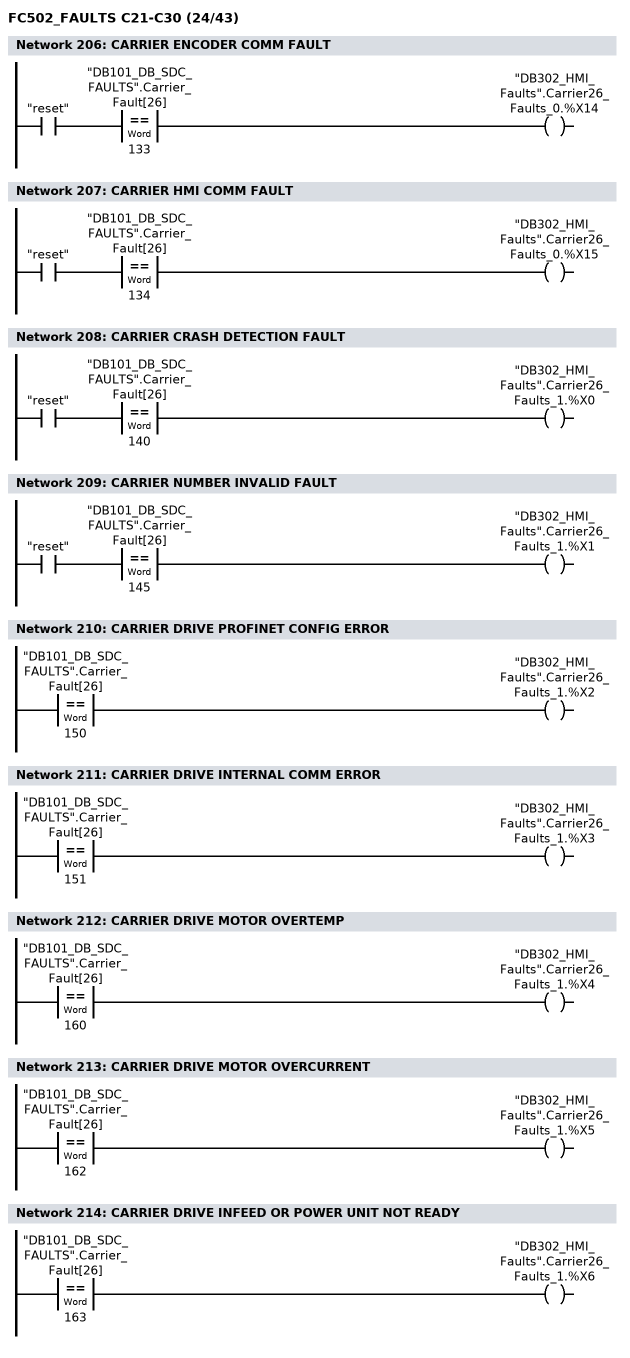
   RUNG wire#powerrail
      Contact( "reset" )
      { S7_Templates := "SrcType := Word" } EQ_Contact(in1 := "DB101_DB_SDC_FAULTS".Carrier_Fault[26], in2 := 133)
      Coil( "DB302_HMI_Faults".Carrier26_Faults_0.%X14 )
   END_RUNG
   // the same network as SCL:
   "DB302_HMI_Faults".Carrier26_Faults_0.%X14 := "reset" AND ("DB101_DB_SDC_FAULTS".Carrier_Fault[26] = 133);
END_REGION

REGION Network 207: CARRIER HMI COMM FAULT
   RUNG wire#powerrail
      Contact( "reset" )
      { S7_Templates := "SrcType := Word" } EQ_Contact(in1 := "DB101_DB_SDC_FAULTS".Carrier_Fault[26], in2 := 134)
      Coil( "DB302_HMI_Faults".Carrier26_Faults_0.%X15 )
   END_RUNG
   // the same network as SCL:
   "DB302_HMI_Faults".Carrier26_Faults_0.%X15 := "reset" AND ("DB101_DB_SDC_FAULTS".Carrier_Fault[26] = 134);
END_REGION

REGION Network 208: CARRIER CRASH DETECTION FAULT
   RUNG wire#powerrail
      Contact( "reset" )
      { S7_Templates := "SrcType := Word" } EQ_Contact(in1 := "DB101_DB_SDC_FAULTS".Carrier_Fault[26], in2 := 140)
      Coil( "DB302_HMI_Faults".Carrier26_Faults_1.%X0 )
   END_RUNG
   // the same network as SCL:
   "DB302_HMI_Faults".Carrier26_Faults_1.%X0 := "reset" AND ("DB101_DB_SDC_FAULTS".Carrier_Fault[26] = 140);
END_REGION

REGION Network 209: CARRIER NUMBER INVALID FAULT
   RUNG wire#powerrail
      Contact( "reset" )
      { S7_Templates := "SrcType := Word" } EQ_Contact(in1 := "DB101_DB_SDC_FAULTS".Carrier_Fault[26], in2 := 145)
      Coil( "DB302_HMI_Faults".Carrier26_Faults_1.%X1 )
   END_RUNG
   // the same network as SCL:
   "DB302_HMI_Faults".Carrier26_Faults_1.%X1 := "reset" AND ("DB101_DB_SDC_FAULTS".Carrier_Fault[26] = 145);
END_REGION

REGION Network 210: CARRIER DRIVE PROFINET CONFIG ERROR
   RUNG wire#powerrail
      { S7_Templates := "SrcType := Word" } EQ_Contact(in1 := "DB101_DB_SDC_FAULTS".Carrier_Fault[26], in2 := 150)
      Coil( "DB302_HMI_Faults".Carrier26_Faults_1.%X2 )
   END_RUNG
   // the same network as SCL:
   "DB302_HMI_Faults".Carrier26_Faults_1.%X2 := "DB101_DB_SDC_FAULTS".Carrier_Fault[26] = 150;
END_REGION

REGION Network 211: CARRIER DRIVE INTERNAL COMM ERROR
   RUNG wire#powerrail
      { S7_Templates := "SrcType := Word" } EQ_Contact(in1 := "DB101_DB_SDC_FAULTS".Carrier_Fault[26], in2 := 151)
      Coil( "DB302_HMI_Faults".Carrier26_Faults_1.%X3 )
   END_RUNG
   // the same network as SCL:
   "DB302_HMI_Faults".Carrier26_Faults_1.%X3 := "DB101_DB_SDC_FAULTS".Carrier_Fault[26] = 151;
END_REGION

REGION Network 212: CARRIER DRIVE MOTOR OVERTEMP
   RUNG wire#powerrail
      { S7_Templates := "SrcType := Word" } EQ_Contact(in1 := "DB101_DB_SDC_FAULTS".Carrier_Fault[26], in2 := 160)
      Coil( "DB302_HMI_Faults".Carrier26_Faults_1.%X4 )
   END_RUNG
   // the same network as SCL:
   "DB302_HMI_Faults".Carrier26_Faults_1.%X4 := "DB101_DB_SDC_FAULTS".Carrier_Fault[26] = 160;
END_REGION

REGION Network 213: CARRIER DRIVE MOTOR OVERCURRENT
   RUNG wire#powerrail
      { S7_Templates := "SrcType := Word" } EQ_Contact(in1 := "DB101_DB_SDC_FAULTS".Carrier_Fault[26], in2 := 162)
      Coil( "DB302_HMI_Faults".Carrier26_Faults_1.%X5 )
   END_RUNG
   // the same network as SCL:
   "DB302_HMI_Faults".Carrier26_Faults_1.%X5 := "DB101_DB_SDC_FAULTS".Carrier_Fault[26] = 162;
END_REGION

REGION Network 214: CARRIER DRIVE INFEED OR POWER UNIT NOT READY
   RUNG wire#powerrail
      { S7_Templates := "SrcType := Word" } EQ_Contact(in1 := "DB101_DB_SDC_FAULTS".Carrier_Fault[26], in2 := 163)
      Coil( "DB302_HMI_Faults".Carrier26_Faults_1.%X6 )
   END_RUNG
   // the same network as SCL:
   "DB302_HMI_Faults".Carrier26_Faults_1.%X6 := "DB101_DB_SDC_FAULTS".Carrier_Fault[26] = 163;
END_REGION

REGION Network 215: CARRIER DRIVE SHORT CIRCUIT / GROUND FAULT DETECTED
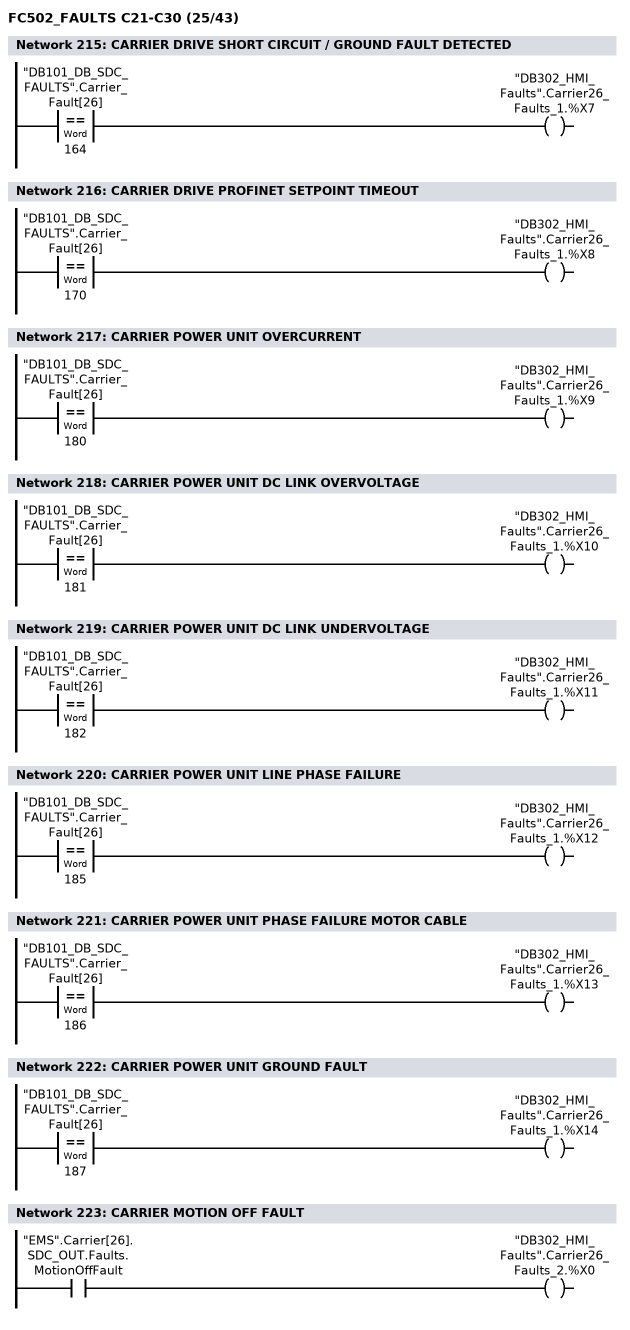
   RUNG wire#powerrail
      { S7_Templates := "SrcType := Word" } EQ_Contact(in1 := "DB101_DB_SDC_FAULTS".Carrier_Fault[26], in2 := 164)
      Coil( "DB302_HMI_Faults".Carrier26_Faults_1.%X7 )
   END_RUNG
   // the same network as SCL:
   "DB302_HMI_Faults".Carrier26_Faults_1.%X7 := "DB101_DB_SDC_FAULTS".Carrier_Fault[26] = 164;
END_REGION

REGION Network 216: CARRIER DRIVE PROFINET SETPOINT TIMEOUT
   RUNG wire#powerrail
      { S7_Templates := "SrcType := Word" } EQ_Contact(in1 := "DB101_DB_SDC_FAULTS".Carrier_Fault[26], in2 := 170)
      Coil( "DB302_HMI_Faults".Carrier26_Faults_1.%X8 )
   END_RUNG
   // the same network as SCL:
   "DB302_HMI_Faults".Carrier26_Faults_1.%X8 := "DB101_DB_SDC_FAULTS".Carrier_Fault[26] = 170;
END_REGION

REGION Network 217: CARRIER POWER UNIT OVERCURRENT
   RUNG wire#powerrail
      { S7_Templates := "SrcType := Word" } EQ_Contact(in1 := "DB101_DB_SDC_FAULTS".Carrier_Fault[26], in2 := 180)
      Coil( "DB302_HMI_Faults".Carrier26_Faults_1.%X9 )
   END_RUNG
   // the same network as SCL:
   "DB302_HMI_Faults".Carrier26_Faults_1.%X9 := "DB101_DB_SDC_FAULTS".Carrier_Fault[26] = 180;
END_REGION

REGION Network 218: CARRIER POWER UNIT DC LINK OVERVOLTAGE
   RUNG wire#powerrail
      { S7_Templates := "SrcType := Word" } EQ_Contact(in1 := "DB101_DB_SDC_FAULTS".Carrier_Fault[26], in2 := 181)
      Coil( "DB302_HMI_Faults".Carrier26_Faults_1.%X10 )
   END_RUNG
   // the same network as SCL:
   "DB302_HMI_Faults".Carrier26_Faults_1.%X10 := "DB101_DB_SDC_FAULTS".Carrier_Fault[26] = 181;
END_REGION

REGION Network 219: CARRIER POWER UNIT DC LINK UNDERVOLTAGE
   RUNG wire#powerrail
      { S7_Templates := "SrcType := Word" } EQ_Contact(in1 := "DB101_DB_SDC_FAULTS".Carrier_Fault[26], in2 := 182)
      Coil( "DB302_HMI_Faults".Carrier26_Faults_1.%X11 )
   END_RUNG
   // the same network as SCL:
   "DB302_HMI_Faults".Carrier26_Faults_1.%X11 := "DB101_DB_SDC_FAULTS".Carrier_Fault[26] = 182;
END_REGION

REGION Network 220: CARRIER POWER UNIT LINE PHASE FAILURE
   RUNG wire#powerrail
      { S7_Templates := "SrcType := Word" } EQ_Contact(in1 := "DB101_DB_SDC_FAULTS".Carrier_Fault[26], in2 := 185)
      Coil( "DB302_HMI_Faults".Carrier26_Faults_1.%X12 )
   END_RUNG
   // the same network as SCL:
   "DB302_HMI_Faults".Carrier26_Faults_1.%X12 := "DB101_DB_SDC_FAULTS".Carrier_Fault[26] = 185;
END_REGION

REGION Network 221: CARRIER POWER UNIT PHASE FAILURE MOTOR CABLE
   RUNG wire#powerrail
      { S7_Templates := "SrcType := Word" } EQ_Contact(in1 := "DB101_DB_SDC_FAULTS".Carrier_Fault[26], in2 := 186)
      Coil( "DB302_HMI_Faults".Carrier26_Faults_1.%X13 )
   END_RUNG
   // the same network as SCL:
   "DB302_HMI_Faults".Carrier26_Faults_1.%X13 := "DB101_DB_SDC_FAULTS".Carrier_Fault[26] = 186;
END_REGION

REGION Network 222: CARRIER POWER UNIT GROUND FAULT
   RUNG wire#powerrail
      { S7_Templates := "SrcType := Word" } EQ_Contact(in1 := "DB101_DB_SDC_FAULTS".Carrier_Fault[26], in2 := 187)
      Coil( "DB302_HMI_Faults".Carrier26_Faults_1.%X14 )
   END_RUNG
   // the same network as SCL:
   "DB302_HMI_Faults".Carrier26_Faults_1.%X14 := "DB101_DB_SDC_FAULTS".Carrier_Fault[26] = 187;
END_REGION

REGION Network 223: CARRIER MOTION OFF FAULT
   RUNG wire#powerrail
      Contact( "EMS".Carrier[26].SDC_OUT.Faults.MotionOffFault )
      Coil( "DB302_HMI_Faults".Carrier26_Faults_2.%X0 )
   END_RUNG
   // the same network as SCL:
   "DB302_HMI_Faults".Carrier26_Faults_2.%X0 := "EMS".Carrier[26].SDC_OUT.Faults.MotionOffFault;
END_REGION

REGION Network 224: CARRIER MOTION ON FAULT
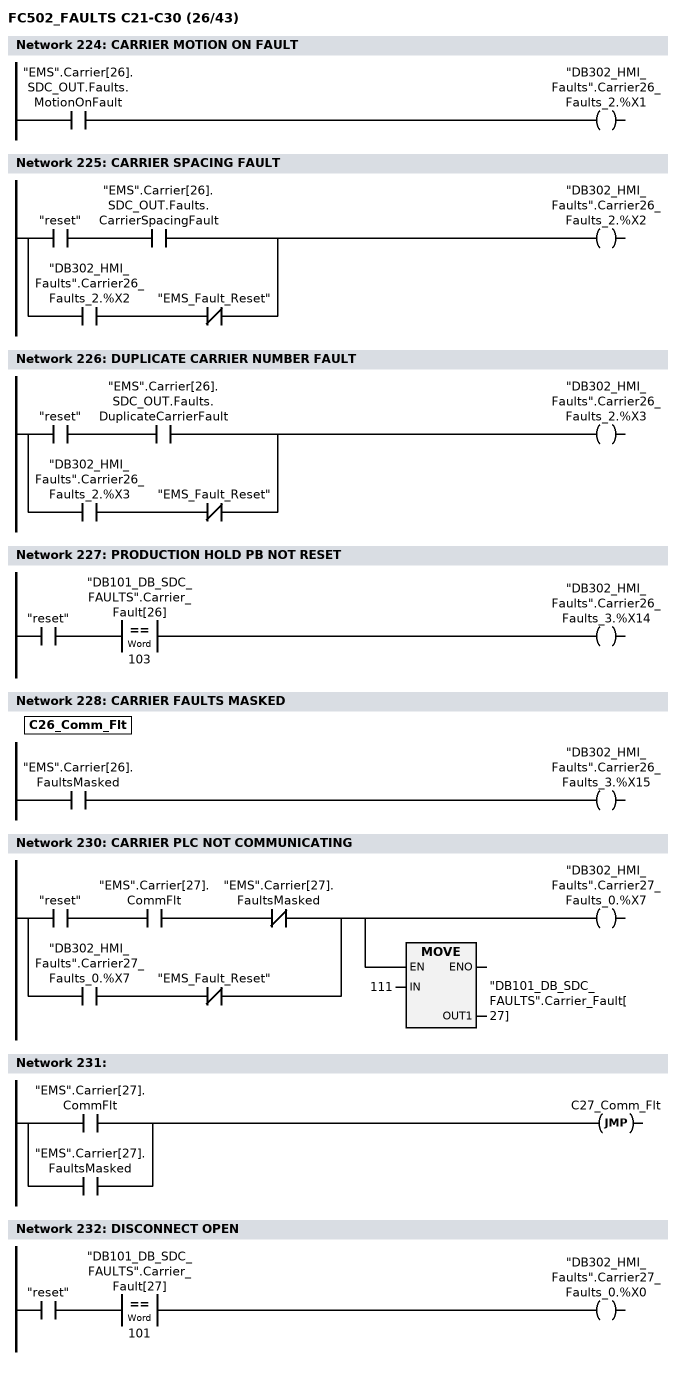
   RUNG wire#powerrail
      Contact( "EMS".Carrier[26].SDC_OUT.Faults.MotionOnFault )
      Coil( "DB302_HMI_Faults".Carrier26_Faults_2.%X1 )
   END_RUNG
   // the same network as SCL:
   "DB302_HMI_Faults".Carrier26_Faults_2.%X1 := "EMS".Carrier[26].SDC_OUT.Faults.MotionOnFault;
END_REGION

REGION Network 225: CARRIER SPACING FAULT
   RUNG wire#powerrail
      Contact( "reset" )
      Contact( "EMS".Carrier[26].SDC_OUT.Faults.CarrierSpacingFault )
      wire#w1
      Coil( "DB302_HMI_Faults".Carrier26_Faults_2.%X2 )
   END_RUNG
   RUNG wire#powerrail
      Contact( "DB302_HMI_Faults".Carrier26_Faults_2.%X2 )
      I_Contact( "EMS_Fault_Reset" )
   END_RUNG wire#w1
   // the same network as SCL:
   "DB302_HMI_Faults".Carrier26_Faults_2.%X2 := ("reset" AND "EMS".Carrier[26].SDC_OUT.Faults.CarrierSpacingFault) OR ("DB302_HMI_Faults".Carrier26_Faults_2.%X2 AND NOT "EMS_Fault_Reset");
END_REGION

REGION Network 226: DUPLICATE CARRIER NUMBER FAULT
   RUNG wire#powerrail
      Contact( "reset" )
      Contact( "EMS".Carrier[26].SDC_OUT.Faults.DuplicateCarrierFault )
      wire#w1
      Coil( "DB302_HMI_Faults".Carrier26_Faults_2.%X3 )
   END_RUNG
   RUNG wire#powerrail
      Contact( "DB302_HMI_Faults".Carrier26_Faults_2.%X3 )
      I_Contact( "EMS_Fault_Reset" )
   END_RUNG wire#w1
   // the same network as SCL:
   "DB302_HMI_Faults".Carrier26_Faults_2.%X3 := ("reset" AND "EMS".Carrier[26].SDC_OUT.Faults.DuplicateCarrierFault) OR ("DB302_HMI_Faults".Carrier26_Faults_2.%X3 AND NOT "EMS_Fault_Reset");
END_REGION

REGION Network 227: PRODUCTION HOLD PB NOT RESET
   RUNG wire#powerrail
      Contact( "reset" )
      { S7_Templates := "SrcType := Word" } EQ_Contact(in1 := "DB101_DB_SDC_FAULTS".Carrier_Fault[26], in2 := 103)
      Coil( "DB302_HMI_Faults".Carrier26_Faults_3.%X14 )
   END_RUNG
   // the same network as SCL:
   "DB302_HMI_Faults".Carrier26_Faults_3.%X14 := "reset" AND ("DB101_DB_SDC_FAULTS".Carrier_Fault[26] = 103);
END_REGION

REGION Network 228: CARRIER FAULTS MASKED
   Label( C26_Comm_Flt )
   RUNG wire#powerrail
      Contact( "EMS".Carrier[26].FaultsMasked )
      Coil( "DB302_HMI_Faults".Carrier26_Faults_3.%X15 )
   END_RUNG
   // the same network as SCL:
   C26_Comm_Flt:
   "DB302_HMI_Faults".Carrier26_Faults_3.%X15 := "EMS".Carrier[26].FaultsMasked;
END_REGION

REGION Network 229: CARRIER 27 FAULTS
END_REGION

REGION Network 230: CARRIER PLC NOT COMMUNICATING
   RUNG wire#powerrail
      Contact( "reset" )
      Contact( "EMS".Carrier[27].CommFlt )
      I_Contact( "EMS".Carrier[27].FaultsMasked )
      wire#w1
      Coil( "DB302_HMI_Faults".Carrier27_Faults_0.%X7 )
   END_RUNG
   RUNG wire#powerrail
      Contact( "DB302_HMI_Faults".Carrier27_Faults_0.%X7 )
      I_Contact( "EMS_Fault_Reset" )
   END_RUNG wire#w1
   RUNG wire#w1
      Move(in := 111, out1 => "DB101_DB_SDC_FAULTS".Carrier_Fault[27])
   END_RUNG
   // the same network as SCL:
   "DB302_HMI_Faults".Carrier27_Faults_0.%X7 := ("reset" AND "EMS".Carrier[27].CommFlt AND NOT "EMS".Carrier[27].FaultsMasked) OR ("DB302_HMI_Faults".Carrier27_Faults_0.%X7 AND NOT "EMS_Fault_Reset");
   IF "DB302_HMI_Faults".Carrier27_Faults_0.%X7 THEN "DB101_DB_SDC_FAULTS".Carrier_Fault[27] := 111; END_IF;
END_REGION

REGION Network 231
   RUNG wire#powerrail
      Contact( "EMS".Carrier[27].CommFlt )
      wire#w1
      JumpCoil( C27_Comm_Flt )
   END_RUNG
   RUNG wire#powerrail
      Contact( "EMS".Carrier[27].FaultsMasked )
   END_RUNG wire#w1
   // the same network as SCL:
   IF "EMS".Carrier[27].CommFlt OR "EMS".Carrier[27].FaultsMasked THEN GOTO C27_Comm_Flt; END_IF;
END_REGION

REGION Network 232: DISCONNECT OPEN
   RUNG wire#powerrail
      Contact( "reset" )
      { S7_Templates := "SrcType := Word" } EQ_Contact(in1 := "DB101_DB_SDC_FAULTS".Carrier_Fault[27], in2 := 101)
      Coil( "DB302_HMI_Faults".Carrier27_Faults_0.%X0 )
   END_RUNG
   // the same network as SCL:
   "DB302_HMI_Faults".Carrier27_Faults_0.%X0 := "reset" AND ("DB101_DB_SDC_FAULTS".Carrier_Fault[27] = 101);
END_REGION

REGION Network 233: PROFINET FAULT
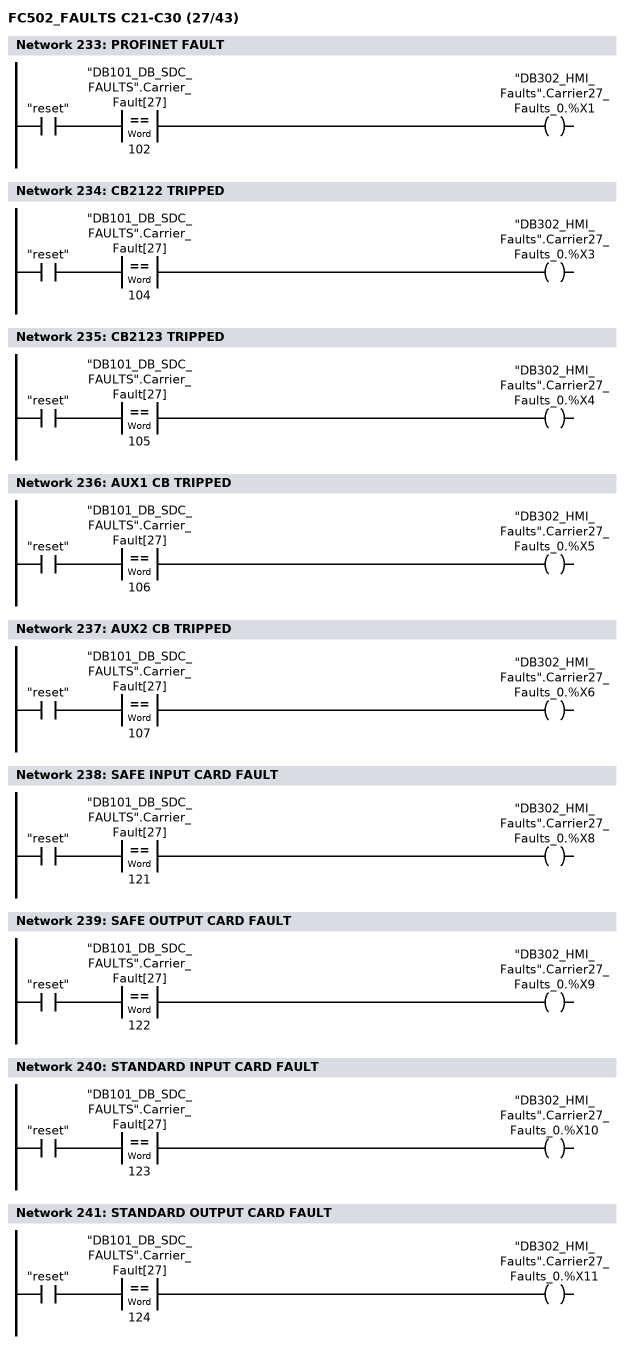
   RUNG wire#powerrail
      Contact( "reset" )
      { S7_Templates := "SrcType := Word" } EQ_Contact(in1 := "DB101_DB_SDC_FAULTS".Carrier_Fault[27], in2 := 102)
      Coil( "DB302_HMI_Faults".Carrier27_Faults_0.%X1 )
   END_RUNG
   // the same network as SCL:
   "DB302_HMI_Faults".Carrier27_Faults_0.%X1 := "reset" AND ("DB101_DB_SDC_FAULTS".Carrier_Fault[27] = 102);
END_REGION

REGION Network 234: CB2122 TRIPPED
   RUNG wire#powerrail
      Contact( "reset" )
      { S7_Templates := "SrcType := Word" } EQ_Contact(in1 := "DB101_DB_SDC_FAULTS".Carrier_Fault[27], in2 := 104)
      Coil( "DB302_HMI_Faults".Carrier27_Faults_0.%X3 )
   END_RUNG
   // the same network as SCL:
   "DB302_HMI_Faults".Carrier27_Faults_0.%X3 := "reset" AND ("DB101_DB_SDC_FAULTS".Carrier_Fault[27] = 104);
END_REGION

REGION Network 235: CB2123 TRIPPED
   RUNG wire#powerrail
      Contact( "reset" )
      { S7_Templates := "SrcType := Word" } EQ_Contact(in1 := "DB101_DB_SDC_FAULTS".Carrier_Fault[27], in2 := 105)
      Coil( "DB302_HMI_Faults".Carrier27_Faults_0.%X4 )
   END_RUNG
   // the same network as SCL:
   "DB302_HMI_Faults".Carrier27_Faults_0.%X4 := "reset" AND ("DB101_DB_SDC_FAULTS".Carrier_Fault[27] = 105);
END_REGION

REGION Network 236: AUX1 CB TRIPPED
   RUNG wire#powerrail
      Contact( "reset" )
      { S7_Templates := "SrcType := Word" } EQ_Contact(in1 := "DB101_DB_SDC_FAULTS".Carrier_Fault[27], in2 := 106)
      Coil( "DB302_HMI_Faults".Carrier27_Faults_0.%X5 )
   END_RUNG
   // the same network as SCL:
   "DB302_HMI_Faults".Carrier27_Faults_0.%X5 := "reset" AND ("DB101_DB_SDC_FAULTS".Carrier_Fault[27] = 106);
END_REGION

REGION Network 237: AUX2 CB TRIPPED
   RUNG wire#powerrail
      Contact( "reset" )
      { S7_Templates := "SrcType := Word" } EQ_Contact(in1 := "DB101_DB_SDC_FAULTS".Carrier_Fault[27], in2 := 107)
      Coil( "DB302_HMI_Faults".Carrier27_Faults_0.%X6 )
   END_RUNG
   // the same network as SCL:
   "DB302_HMI_Faults".Carrier27_Faults_0.%X6 := "reset" AND ("DB101_DB_SDC_FAULTS".Carrier_Fault[27] = 107);
END_REGION

REGION Network 238: SAFE INPUT CARD FAULT
   RUNG wire#powerrail
      Contact( "reset" )
      { S7_Templates := "SrcType := Word" } EQ_Contact(in1 := "DB101_DB_SDC_FAULTS".Carrier_Fault[27], in2 := 121)
      Coil( "DB302_HMI_Faults".Carrier27_Faults_0.%X8 )
   END_RUNG
   // the same network as SCL:
   "DB302_HMI_Faults".Carrier27_Faults_0.%X8 := "reset" AND ("DB101_DB_SDC_FAULTS".Carrier_Fault[27] = 121);
END_REGION

REGION Network 239: SAFE OUTPUT CARD FAULT
   RUNG wire#powerrail
      Contact( "reset" )
      { S7_Templates := "SrcType := Word" } EQ_Contact(in1 := "DB101_DB_SDC_FAULTS".Carrier_Fault[27], in2 := 122)
      Coil( "DB302_HMI_Faults".Carrier27_Faults_0.%X9 )
   END_RUNG
   // the same network as SCL:
   "DB302_HMI_Faults".Carrier27_Faults_0.%X9 := "reset" AND ("DB101_DB_SDC_FAULTS".Carrier_Fault[27] = 122);
END_REGION

REGION Network 240: STANDARD INPUT CARD FAULT
   RUNG wire#powerrail
      Contact( "reset" )
      { S7_Templates := "SrcType := Word" } EQ_Contact(in1 := "DB101_DB_SDC_FAULTS".Carrier_Fault[27], in2 := 123)
      Coil( "DB302_HMI_Faults".Carrier27_Faults_0.%X10 )
   END_RUNG
   // the same network as SCL:
   "DB302_HMI_Faults".Carrier27_Faults_0.%X10 := "reset" AND ("DB101_DB_SDC_FAULTS".Carrier_Fault[27] = 123);
END_REGION

REGION Network 241: STANDARD OUTPUT CARD FAULT
   RUNG wire#powerrail
      Contact( "reset" )
      { S7_Templates := "SrcType := Word" } EQ_Contact(in1 := "DB101_DB_SDC_FAULTS".Carrier_Fault[27], in2 := 124)
      Coil( "DB302_HMI_Faults".Carrier27_Faults_0.%X11 )
   END_RUNG
   // the same network as SCL:
   "DB302_HMI_Faults".Carrier27_Faults_0.%X11 := "reset" AND ("DB101_DB_SDC_FAULTS".Carrier_Fault[27] = 124);
END_REGION

REGION Network 242: CARRIER ENCODER POSITION FAULT
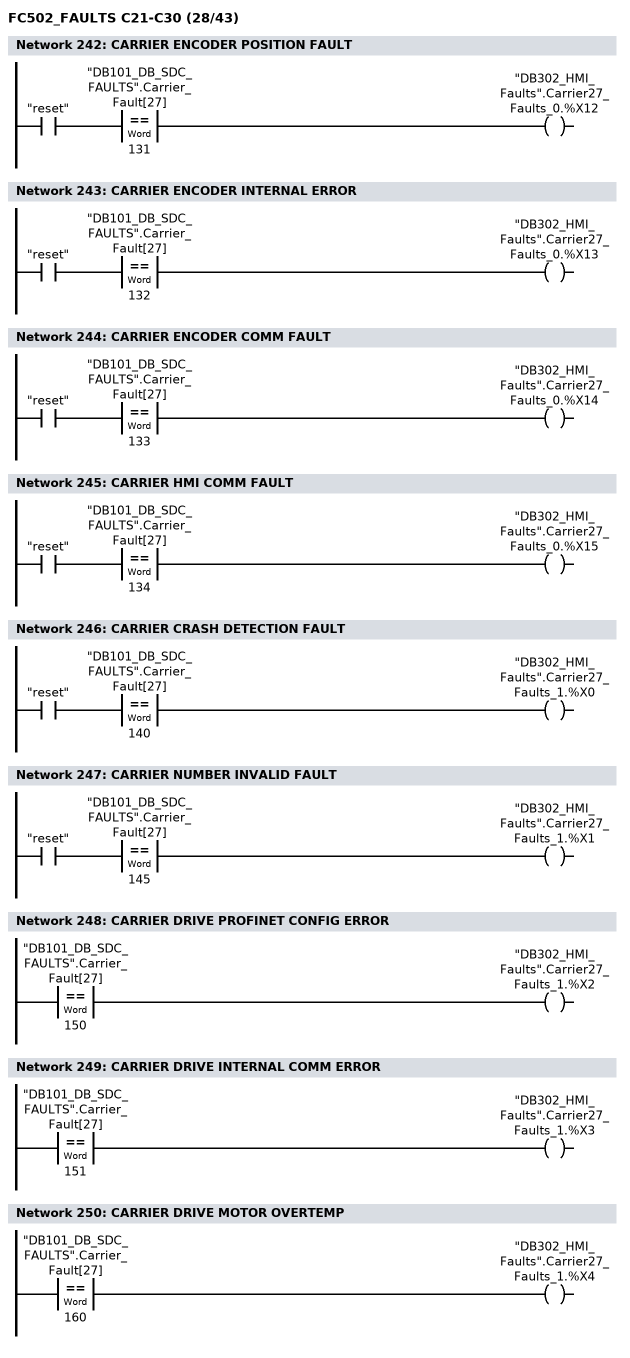
   RUNG wire#powerrail
      Contact( "reset" )
      { S7_Templates := "SrcType := Word" } EQ_Contact(in1 := "DB101_DB_SDC_FAULTS".Carrier_Fault[27], in2 := 131)
      Coil( "DB302_HMI_Faults".Carrier27_Faults_0.%X12 )
   END_RUNG
   // the same network as SCL:
   "DB302_HMI_Faults".Carrier27_Faults_0.%X12 := "reset" AND ("DB101_DB_SDC_FAULTS".Carrier_Fault[27] = 131);
END_REGION

REGION Network 243: CARRIER ENCODER INTERNAL ERROR
   RUNG wire#powerrail
      Contact( "reset" )
      { S7_Templates := "SrcType := Word" } EQ_Contact(in1 := "DB101_DB_SDC_FAULTS".Carrier_Fault[27], in2 := 132)
      Coil( "DB302_HMI_Faults".Carrier27_Faults_0.%X13 )
   END_RUNG
   // the same network as SCL:
   "DB302_HMI_Faults".Carrier27_Faults_0.%X13 := "reset" AND ("DB101_DB_SDC_FAULTS".Carrier_Fault[27] = 132);
END_REGION

REGION Network 244: CARRIER ENCODER COMM FAULT
   RUNG wire#powerrail
      Contact( "reset" )
      { S7_Templates := "SrcType := Word" } EQ_Contact(in1 := "DB101_DB_SDC_FAULTS".Carrier_Fault[27], in2 := 133)
      Coil( "DB302_HMI_Faults".Carrier27_Faults_0.%X14 )
   END_RUNG
   // the same network as SCL:
   "DB302_HMI_Faults".Carrier27_Faults_0.%X14 := "reset" AND ("DB101_DB_SDC_FAULTS".Carrier_Fault[27] = 133);
END_REGION

REGION Network 245: CARRIER HMI COMM FAULT
   RUNG wire#powerrail
      Contact( "reset" )
      { S7_Templates := "SrcType := Word" } EQ_Contact(in1 := "DB101_DB_SDC_FAULTS".Carrier_Fault[27], in2 := 134)
      Coil( "DB302_HMI_Faults".Carrier27_Faults_0.%X15 )
   END_RUNG
   // the same network as SCL:
   "DB302_HMI_Faults".Carrier27_Faults_0.%X15 := "reset" AND ("DB101_DB_SDC_FAULTS".Carrier_Fault[27] = 134);
END_REGION

REGION Network 246: CARRIER CRASH DETECTION FAULT
   RUNG wire#powerrail
      Contact( "reset" )
      { S7_Templates := "SrcType := Word" } EQ_Contact(in1 := "DB101_DB_SDC_FAULTS".Carrier_Fault[27], in2 := 140)
      Coil( "DB302_HMI_Faults".Carrier27_Faults_1.%X0 )
   END_RUNG
   // the same network as SCL:
   "DB302_HMI_Faults".Carrier27_Faults_1.%X0 := "reset" AND ("DB101_DB_SDC_FAULTS".Carrier_Fault[27] = 140);
END_REGION

REGION Network 247: CARRIER NUMBER INVALID FAULT
   RUNG wire#powerrail
      Contact( "reset" )
      { S7_Templates := "SrcType := Word" } EQ_Contact(in1 := "DB101_DB_SDC_FAULTS".Carrier_Fault[27], in2 := 145)
      Coil( "DB302_HMI_Faults".Carrier27_Faults_1.%X1 )
   END_RUNG
   // the same network as SCL:
   "DB302_HMI_Faults".Carrier27_Faults_1.%X1 := "reset" AND ("DB101_DB_SDC_FAULTS".Carrier_Fault[27] = 145);
END_REGION

REGION Network 248: CARRIER DRIVE PROFINET CONFIG ERROR
   RUNG wire#powerrail
      { S7_Templates := "SrcType := Word" } EQ_Contact(in1 := "DB101_DB_SDC_FAULTS".Carrier_Fault[27], in2 := 150)
      Coil( "DB302_HMI_Faults".Carrier27_Faults_1.%X2 )
   END_RUNG
   // the same network as SCL:
   "DB302_HMI_Faults".Carrier27_Faults_1.%X2 := "DB101_DB_SDC_FAULTS".Carrier_Fault[27] = 150;
END_REGION

REGION Network 249: CARRIER DRIVE INTERNAL COMM ERROR
   RUNG wire#powerrail
      { S7_Templates := "SrcType := Word" } EQ_Contact(in1 := "DB101_DB_SDC_FAULTS".Carrier_Fault[27], in2 := 151)
      Coil( "DB302_HMI_Faults".Carrier27_Faults_1.%X3 )
   END_RUNG
   // the same network as SCL:
   "DB302_HMI_Faults".Carrier27_Faults_1.%X3 := "DB101_DB_SDC_FAULTS".Carrier_Fault[27] = 151;
END_REGION

REGION Network 250: CARRIER DRIVE MOTOR OVERTEMP
   RUNG wire#powerrail
      { S7_Templates := "SrcType := Word" } EQ_Contact(in1 := "DB101_DB_SDC_FAULTS".Carrier_Fault[27], in2 := 160)
      Coil( "DB302_HMI_Faults".Carrier27_Faults_1.%X4 )
   END_RUNG
   // the same network as SCL:
   "DB302_HMI_Faults".Carrier27_Faults_1.%X4 := "DB101_DB_SDC_FAULTS".Carrier_Fault[27] = 160;
END_REGION

REGION Network 251: CARRIER DRIVE MOTOR OVERCURRENT
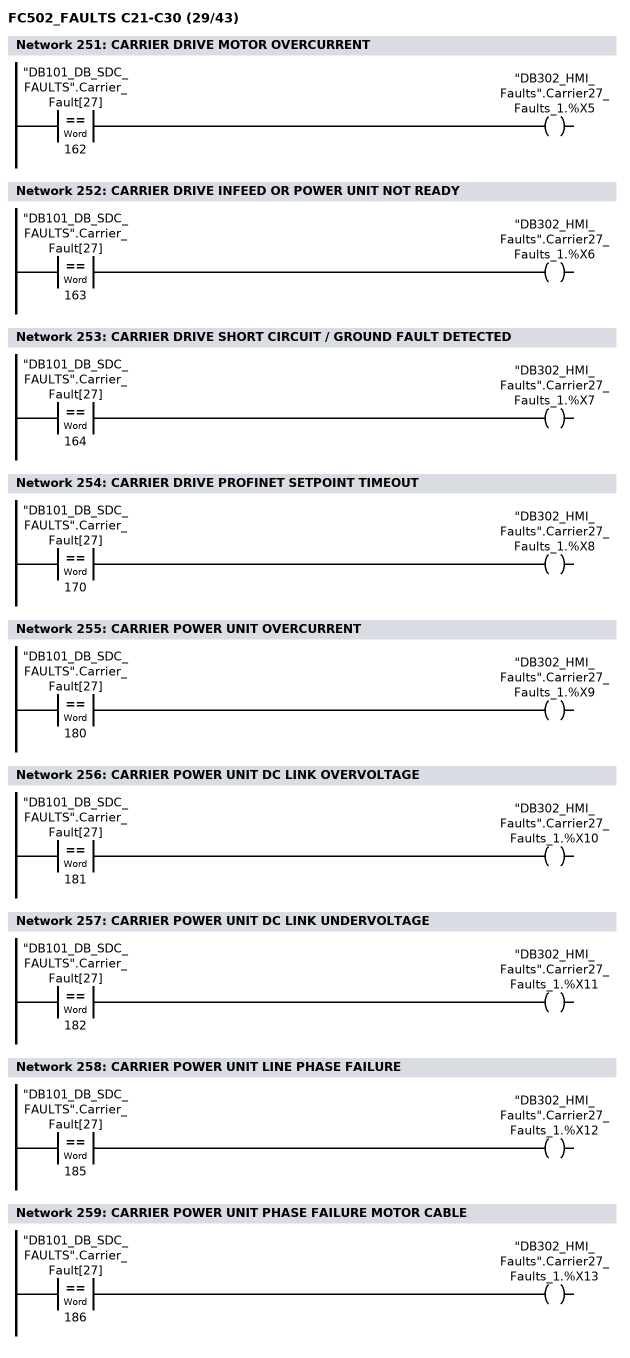
   RUNG wire#powerrail
      { S7_Templates := "SrcType := Word" } EQ_Contact(in1 := "DB101_DB_SDC_FAULTS".Carrier_Fault[27], in2 := 162)
      Coil( "DB302_HMI_Faults".Carrier27_Faults_1.%X5 )
   END_RUNG
   // the same network as SCL:
   "DB302_HMI_Faults".Carrier27_Faults_1.%X5 := "DB101_DB_SDC_FAULTS".Carrier_Fault[27] = 162;
END_REGION

REGION Network 252: CARRIER DRIVE INFEED OR POWER UNIT NOT READY
   RUNG wire#powerrail
      { S7_Templates := "SrcType := Word" } EQ_Contact(in1 := "DB101_DB_SDC_FAULTS".Carrier_Fault[27], in2 := 163)
      Coil( "DB302_HMI_Faults".Carrier27_Faults_1.%X6 )
   END_RUNG
   // the same network as SCL:
   "DB302_HMI_Faults".Carrier27_Faults_1.%X6 := "DB101_DB_SDC_FAULTS".Carrier_Fault[27] = 163;
END_REGION

REGION Network 253: CARRIER DRIVE SHORT CIRCUIT / GROUND FAULT DETECTED
   RUNG wire#powerrail
      { S7_Templates := "SrcType := Word" } EQ_Contact(in1 := "DB101_DB_SDC_FAULTS".Carrier_Fault[27], in2 := 164)
      Coil( "DB302_HMI_Faults".Carrier27_Faults_1.%X7 )
   END_RUNG
   // the same network as SCL:
   "DB302_HMI_Faults".Carrier27_Faults_1.%X7 := "DB101_DB_SDC_FAULTS".Carrier_Fault[27] = 164;
END_REGION

REGION Network 254: CARRIER DRIVE PROFINET SETPOINT TIMEOUT
   RUNG wire#powerrail
      { S7_Templates := "SrcType := Word" } EQ_Contact(in1 := "DB101_DB_SDC_FAULTS".Carrier_Fault[27], in2 := 170)
      Coil( "DB302_HMI_Faults".Carrier27_Faults_1.%X8 )
   END_RUNG
   // the same network as SCL:
   "DB302_HMI_Faults".Carrier27_Faults_1.%X8 := "DB101_DB_SDC_FAULTS".Carrier_Fault[27] = 170;
END_REGION

REGION Network 255: CARRIER POWER UNIT OVERCURRENT
   RUNG wire#powerrail
      { S7_Templates := "SrcType := Word" } EQ_Contact(in1 := "DB101_DB_SDC_FAULTS".Carrier_Fault[27], in2 := 180)
      Coil( "DB302_HMI_Faults".Carrier27_Faults_1.%X9 )
   END_RUNG
   // the same network as SCL:
   "DB302_HMI_Faults".Carrier27_Faults_1.%X9 := "DB101_DB_SDC_FAULTS".Carrier_Fault[27] = 180;
END_REGION

REGION Network 256: CARRIER POWER UNIT DC LINK OVERVOLTAGE
   RUNG wire#powerrail
      { S7_Templates := "SrcType := Word" } EQ_Contact(in1 := "DB101_DB_SDC_FAULTS".Carrier_Fault[27], in2 := 181)
      Coil( "DB302_HMI_Faults".Carrier27_Faults_1.%X10 )
   END_RUNG
   // the same network as SCL:
   "DB302_HMI_Faults".Carrier27_Faults_1.%X10 := "DB101_DB_SDC_FAULTS".Carrier_Fault[27] = 181;
END_REGION

REGION Network 257: CARRIER POWER UNIT DC LINK UNDERVOLTAGE
   RUNG wire#powerrail
      { S7_Templates := "SrcType := Word" } EQ_Contact(in1 := "DB101_DB_SDC_FAULTS".Carrier_Fault[27], in2 := 182)
      Coil( "DB302_HMI_Faults".Carrier27_Faults_1.%X11 )
   END_RUNG
   // the same network as SCL:
   "DB302_HMI_Faults".Carrier27_Faults_1.%X11 := "DB101_DB_SDC_FAULTS".Carrier_Fault[27] = 182;
END_REGION

REGION Network 258: CARRIER POWER UNIT LINE PHASE FAILURE
   RUNG wire#powerrail
      { S7_Templates := "SrcType := Word" } EQ_Contact(in1 := "DB101_DB_SDC_FAULTS".Carrier_Fault[27], in2 := 185)
      Coil( "DB302_HMI_Faults".Carrier27_Faults_1.%X12 )
   END_RUNG
   // the same network as SCL:
   "DB302_HMI_Faults".Carrier27_Faults_1.%X12 := "DB101_DB_SDC_FAULTS".Carrier_Fault[27] = 185;
END_REGION

REGION Network 259: CARRIER POWER UNIT PHASE FAILURE MOTOR CABLE
   RUNG wire#powerrail
      { S7_Templates := "SrcType := Word" } EQ_Contact(in1 := "DB101_DB_SDC_FAULTS".Carrier_Fault[27], in2 := 186)
      Coil( "DB302_HMI_Faults".Carrier27_Faults_1.%X13 )
   END_RUNG
   // the same network as SCL:
   "DB302_HMI_Faults".Carrier27_Faults_1.%X13 := "DB101_DB_SDC_FAULTS".Carrier_Fault[27] = 186;
END_REGION

REGION Network 260: CARRIER POWER UNIT GROUND FAULT
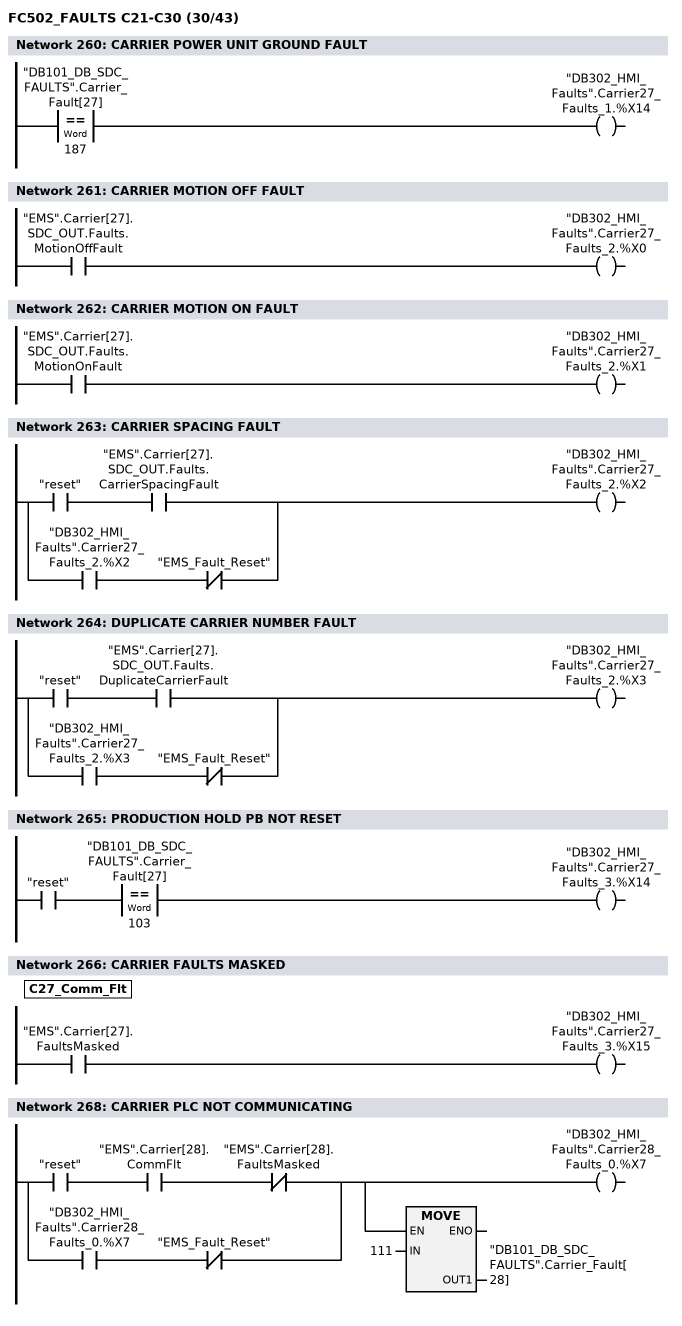
   RUNG wire#powerrail
      { S7_Templates := "SrcType := Word" } EQ_Contact(in1 := "DB101_DB_SDC_FAULTS".Carrier_Fault[27], in2 := 187)
      Coil( "DB302_HMI_Faults".Carrier27_Faults_1.%X14 )
   END_RUNG
   // the same network as SCL:
   "DB302_HMI_Faults".Carrier27_Faults_1.%X14 := "DB101_DB_SDC_FAULTS".Carrier_Fault[27] = 187;
END_REGION

REGION Network 261: CARRIER MOTION OFF FAULT
   RUNG wire#powerrail
      Contact( "EMS".Carrier[27].SDC_OUT.Faults.MotionOffFault )
      Coil( "DB302_HMI_Faults".Carrier27_Faults_2.%X0 )
   END_RUNG
   // the same network as SCL:
   "DB302_HMI_Faults".Carrier27_Faults_2.%X0 := "EMS".Carrier[27].SDC_OUT.Faults.MotionOffFault;
END_REGION

REGION Network 262: CARRIER MOTION ON FAULT
   RUNG wire#powerrail
      Contact( "EMS".Carrier[27].SDC_OUT.Faults.MotionOnFault )
      Coil( "DB302_HMI_Faults".Carrier27_Faults_2.%X1 )
   END_RUNG
   // the same network as SCL:
   "DB302_HMI_Faults".Carrier27_Faults_2.%X1 := "EMS".Carrier[27].SDC_OUT.Faults.MotionOnFault;
END_REGION

REGION Network 263: CARRIER SPACING FAULT
   RUNG wire#powerrail
      Contact( "reset" )
      Contact( "EMS".Carrier[27].SDC_OUT.Faults.CarrierSpacingFault )
      wire#w1
      Coil( "DB302_HMI_Faults".Carrier27_Faults_2.%X2 )
   END_RUNG
   RUNG wire#powerrail
      Contact( "DB302_HMI_Faults".Carrier27_Faults_2.%X2 )
      I_Contact( "EMS_Fault_Reset" )
   END_RUNG wire#w1
   // the same network as SCL:
   "DB302_HMI_Faults".Carrier27_Faults_2.%X2 := ("reset" AND "EMS".Carrier[27].SDC_OUT.Faults.CarrierSpacingFault) OR ("DB302_HMI_Faults".Carrier27_Faults_2.%X2 AND NOT "EMS_Fault_Reset");
END_REGION

REGION Network 264: DUPLICATE CARRIER NUMBER FAULT
   RUNG wire#powerrail
      Contact( "reset" )
      Contact( "EMS".Carrier[27].SDC_OUT.Faults.DuplicateCarrierFault )
      wire#w1
      Coil( "DB302_HMI_Faults".Carrier27_Faults_2.%X3 )
   END_RUNG
   RUNG wire#powerrail
      Contact( "DB302_HMI_Faults".Carrier27_Faults_2.%X3 )
      I_Contact( "EMS_Fault_Reset" )
   END_RUNG wire#w1
   // the same network as SCL:
   "DB302_HMI_Faults".Carrier27_Faults_2.%X3 := ("reset" AND "EMS".Carrier[27].SDC_OUT.Faults.DuplicateCarrierFault) OR ("DB302_HMI_Faults".Carrier27_Faults_2.%X3 AND NOT "EMS_Fault_Reset");
END_REGION

REGION Network 265: PRODUCTION HOLD PB NOT RESET
   RUNG wire#powerrail
      Contact( "reset" )
      { S7_Templates := "SrcType := Word" } EQ_Contact(in1 := "DB101_DB_SDC_FAULTS".Carrier_Fault[27], in2 := 103)
      Coil( "DB302_HMI_Faults".Carrier27_Faults_3.%X14 )
   END_RUNG
   // the same network as SCL:
   "DB302_HMI_Faults".Carrier27_Faults_3.%X14 := "reset" AND ("DB101_DB_SDC_FAULTS".Carrier_Fault[27] = 103);
END_REGION

REGION Network 266: CARRIER FAULTS MASKED
   Label( C27_Comm_Flt )
   RUNG wire#powerrail
      Contact( "EMS".Carrier[27].FaultsMasked )
      Coil( "DB302_HMI_Faults".Carrier27_Faults_3.%X15 )
   END_RUNG
   // the same network as SCL:
   C27_Comm_Flt:
   "DB302_HMI_Faults".Carrier27_Faults_3.%X15 := "EMS".Carrier[27].FaultsMasked;
END_REGION

REGION Network 267: CARRIER 28 FAULTS
END_REGION

REGION Network 268: CARRIER PLC NOT COMMUNICATING
   RUNG wire#powerrail
      Contact( "reset" )
      Contact( "EMS".Carrier[28].CommFlt )
      I_Contact( "EMS".Carrier[28].FaultsMasked )
      wire#w1
      Coil( "DB302_HMI_Faults".Carrier28_Faults_0.%X7 )
   END_RUNG
   RUNG wire#powerrail
      Contact( "DB302_HMI_Faults".Carrier28_Faults_0.%X7 )
      I_Contact( "EMS_Fault_Reset" )
   END_RUNG wire#w1
   RUNG wire#w1
      Move(in := 111, out1 => "DB101_DB_SDC_FAULTS".Carrier_Fault[28])
   END_RUNG
   // the same network as SCL:
   "DB302_HMI_Faults".Carrier28_Faults_0.%X7 := ("reset" AND "EMS".Carrier[28].CommFlt AND NOT "EMS".Carrier[28].FaultsMasked) OR ("DB302_HMI_Faults".Carrier28_Faults_0.%X7 AND NOT "EMS_Fault_Reset");
   IF "DB302_HMI_Faults".Carrier28_Faults_0.%X7 THEN "DB101_DB_SDC_FAULTS".Carrier_Fault[28] := 111; END_IF;
END_REGION

REGION Network 269
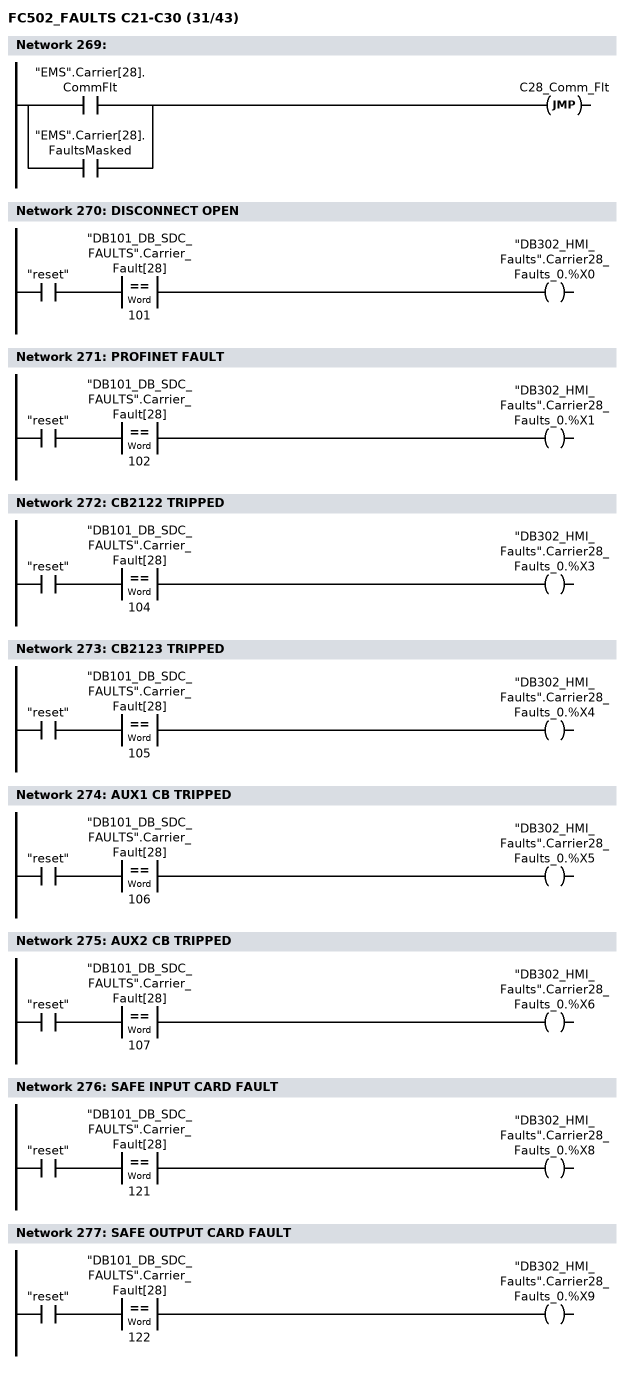
   RUNG wire#powerrail
      Contact( "EMS".Carrier[28].CommFlt )
      wire#w1
      JumpCoil( C28_Comm_Flt )
   END_RUNG
   RUNG wire#powerrail
      Contact( "EMS".Carrier[28].FaultsMasked )
   END_RUNG wire#w1
   // the same network as SCL:
   IF "EMS".Carrier[28].CommFlt OR "EMS".Carrier[28].FaultsMasked THEN GOTO C28_Comm_Flt; END_IF;
END_REGION

REGION Network 270: DISCONNECT OPEN
   RUNG wire#powerrail
      Contact( "reset" )
      { S7_Templates := "SrcType := Word" } EQ_Contact(in1 := "DB101_DB_SDC_FAULTS".Carrier_Fault[28], in2 := 101)
      Coil( "DB302_HMI_Faults".Carrier28_Faults_0.%X0 )
   END_RUNG
   // the same network as SCL:
   "DB302_HMI_Faults".Carrier28_Faults_0.%X0 := "reset" AND ("DB101_DB_SDC_FAULTS".Carrier_Fault[28] = 101);
END_REGION

REGION Network 271: PROFINET FAULT
   RUNG wire#powerrail
      Contact( "reset" )
      { S7_Templates := "SrcType := Word" } EQ_Contact(in1 := "DB101_DB_SDC_FAULTS".Carrier_Fault[28], in2 := 102)
      Coil( "DB302_HMI_Faults".Carrier28_Faults_0.%X1 )
   END_RUNG
   // the same network as SCL:
   "DB302_HMI_Faults".Carrier28_Faults_0.%X1 := "reset" AND ("DB101_DB_SDC_FAULTS".Carrier_Fault[28] = 102);
END_REGION

REGION Network 272: CB2122 TRIPPED
   RUNG wire#powerrail
      Contact( "reset" )
      { S7_Templates := "SrcType := Word" } EQ_Contact(in1 := "DB101_DB_SDC_FAULTS".Carrier_Fault[28], in2 := 104)
      Coil( "DB302_HMI_Faults".Carrier28_Faults_0.%X3 )
   END_RUNG
   // the same network as SCL:
   "DB302_HMI_Faults".Carrier28_Faults_0.%X3 := "reset" AND ("DB101_DB_SDC_FAULTS".Carrier_Fault[28] = 104);
END_REGION

REGION Network 273: CB2123 TRIPPED
   RUNG wire#powerrail
      Contact( "reset" )
      { S7_Templates := "SrcType := Word" } EQ_Contact(in1 := "DB101_DB_SDC_FAULTS".Carrier_Fault[28], in2 := 105)
      Coil( "DB302_HMI_Faults".Carrier28_Faults_0.%X4 )
   END_RUNG
   // the same network as SCL:
   "DB302_HMI_Faults".Carrier28_Faults_0.%X4 := "reset" AND ("DB101_DB_SDC_FAULTS".Carrier_Fault[28] = 105);
END_REGION

REGION Network 274: AUX1 CB TRIPPED
   RUNG wire#powerrail
      Contact( "reset" )
      { S7_Templates := "SrcType := Word" } EQ_Contact(in1 := "DB101_DB_SDC_FAULTS".Carrier_Fault[28], in2 := 106)
      Coil( "DB302_HMI_Faults".Carrier28_Faults_0.%X5 )
   END_RUNG
   // the same network as SCL:
   "DB302_HMI_Faults".Carrier28_Faults_0.%X5 := "reset" AND ("DB101_DB_SDC_FAULTS".Carrier_Fault[28] = 106);
END_REGION

REGION Network 275: AUX2 CB TRIPPED
   RUNG wire#powerrail
      Contact( "reset" )
      { S7_Templates := "SrcType := Word" } EQ_Contact(in1 := "DB101_DB_SDC_FAULTS".Carrier_Fault[28], in2 := 107)
      Coil( "DB302_HMI_Faults".Carrier28_Faults_0.%X6 )
   END_RUNG
   // the same network as SCL:
   "DB302_HMI_Faults".Carrier28_Faults_0.%X6 := "reset" AND ("DB101_DB_SDC_FAULTS".Carrier_Fault[28] = 107);
END_REGION

REGION Network 276: SAFE INPUT CARD FAULT
   RUNG wire#powerrail
      Contact( "reset" )
      { S7_Templates := "SrcType := Word" } EQ_Contact(in1 := "DB101_DB_SDC_FAULTS".Carrier_Fault[28], in2 := 121)
      Coil( "DB302_HMI_Faults".Carrier28_Faults_0.%X8 )
   END_RUNG
   // the same network as SCL:
   "DB302_HMI_Faults".Carrier28_Faults_0.%X8 := "reset" AND ("DB101_DB_SDC_FAULTS".Carrier_Fault[28] = 121);
END_REGION
